// TIA Portal project "CHM_BORDEIRA_20190721" (V15) (continued)
DATA_BLOCK "62_Warning_Data"   // DB62
{ S7_Optimized_Access := 'FALSE' }
VERSION : 0.1
   VAR
      IGG_WARNING_WORD_01 : Word;
      IGG_WARNING_WORD_02 : Word;
      IGG_WARNING_WORD_03 : Word;
      IGG_WARNING_WORD_04 : Word;
      IGG_WARNING_WORD_05 : Word;
      IGG_WARNING_WORD_06 : Word;
      IGG_WARNING_WORD_07 : Word;
      IGG_WARNING_WORD_08 : Word;
      WRNG_PRSNT : Bool;
   END_VAR
BEGIN
END_DATA_BLOCK

DATA_BLOCK "63_E500 Fuel Pumps Not Working_DB"   // DB63
{ S7_Optimized_Access := 'TRUE' }
VERSION : 0.1
// stored: InstanceOfName 63_E500 Fuel Pumps Not Working
"63_E500 Fuel Pumps Not Working"
BEGIN
END_DATA_BLOCK

DATA_BLOCK "64_Message_Data"   // DB64
{ S7_Optimized_Access := 'FALSE' }
VERSION : 0.1
   VAR
      IGG_MESSAGE_WORD_01 : Word;
      IGG_MESSAGE_WORD_02 : Word;
      IGG_MESSAGE_WORD_03 : Word;
      IGG_MESSAGE_WORD_04 : Word;
      IGG_MESSAGE_WORD_05 : Word;
      IGG_MESSAGE_WORD_06 : Word;
      IGG_MESSAGE_WORD_07 : Word;
      IGG_MESSAGE_WORD_08 : Word;
      MSG_PRSNT : Bool;
   END_VAR
BEGIN
END_DATA_BLOCK

DATA_BLOCK "63_Safety System Interlock_IDB"   // DB65
{ S7_Optimized_Access := 'TRUE' }
VERSION : 0.1
// stored: InstanceOfName 64_Safety System Interlock
"64_Safety System Interlock"
BEGIN
END_DATA_BLOCK

DATA_BLOCK "66_Event_Data"   // DB66
{ S7_Optimized_Access := 'FALSE' }
VERSION : 0.1
   VAR
      IGG_EVENT_WORD_01 : Word;
      IGG_EVENT_WORD_02 : Word;
      IGG_EVENT_WORD_03 : Word;
      IGG_EVENT_WORD_04 : Word;
      IGG_EVENT_WORD_05 : Word;
      IGG_EVENT_WORD_06 : Word;
      IGG_EVENT_WORD_07 : Word;
      IGG_EVENT_WORD_08 : Word;
      EVENT_PRSNT : Bool;
   END_VAR
BEGIN
END_DATA_BLOCK

DATA_BLOCK "Alarms_Acknowledge"   // DB67
{ S7_Optimized_Access := 'FALSE' }
VERSION : 0.1
   VAR
      IGG_ALARM_ACKNLG_1 : Word;
      IGG_ALARM_ACKNLG_2 : Word;
      IGG_ALARM_ACKNLG_3 : Word;
      IGG_ALARM_ACKNLG_4 : Word;
      IGG_ALARM_ACKNLG_5 : Word;
      IGG_ALARM_ACKNLG_6 : Word;
   END_VAR
BEGIN
END_DATA_BLOCK

DATA_BLOCK "68_Sys_Status_Data"   // DB68
TITLE = System Status Data
{ S7_Optimized_Access := 'TRUE' }
AUTHOR : JRS
VERSION : 0.1
// Data area for system status information as required by the code
   VAR
      VLVS_AT_INIT : Bool;   // All valves at initial position
      INTRLKS_OK : Bool;   // System interlocks ok
      IA_PRES_IN_RNG : Bool;   // IA Pressure Within Range - PIT112
      CSW_IL_PRES_IN_RNG : Bool;   // CSW Inlet pressure within range - PIT359
      FUEL_PRES_IN_RNG : Bool;   // Fuel pressure within range - PIT204
      OP_PRES_IN_RNG : Bool;   // Output pressure within range - PIT402
      CRG_BLNK_MODE : Bool;   // 1 = Cargon blanketing mode, 0 = Not
      "LOG IGG" : Bool;   // Tag for logging IGG signals
      "STOP LOG IGG" : Bool;
      "LOG IGG Simulator" : Bool;
      "TRUE for HMI" : Bool;
      "E139_SET_SPEED Aux" : Real;
      "E139_SET_SPEED Aux Bool" : Bool;
      "CSW OVR Stop Latched" : Bool;
      "CSW Puls" : Bool;
      "STL Puls" : Bool;
   END_VAR
BEGIN
END_DATA_BLOCK

DATA_BLOCK "503_WARNING CHCK_IDB"   // DB69
{ S7_Optimized_Access := 'TRUE' }
VERSION : 0.1
// stored: InstanceOfName 503_ALARM CHCK
"503_ALARM CHCK"
BEGIN
END_DATA_BLOCK

DATA_BLOCK "CSW_Animation_DB"   // DB71
{ S7_Optimized_Access := 'TRUE' }
VERSION : 0.1
// stored: InstanceOfName Animation
"Animation"
BEGIN
END_DATA_BLOCK

DATA_BLOCK "Ful Pump Ani Animation_DB"   // DB72
{ S7_Optimized_Access := 'TRUE' }
VERSION : 0.1
// stored: InstanceOfName Animation
"Animation"
BEGIN
END_DATA_BLOCK

DATA_BLOCK "IDB_E139"   // DB139
{ S7_Optimized_Access := 'TRUE' }
VERSION : 0.1
// stored: InstanceOfName Animation
"Animation"
BEGIN
END_DATA_BLOCK

DATA_BLOCK "IDB_E500A_Animation"   // DB500
{ S7_Optimized_Access := 'TRUE' }
VERSION : 0.1
// stored: InstanceOfName Animation
"Animation"
BEGIN
END_DATA_BLOCK

DATA_BLOCK "IDB_E500B_Animation"   // DB501
{ S7_Optimized_Access := 'TRUE' }
VERSION : 0.1
// stored: InstanceOfName Animation
"Animation"
BEGIN
END_DATA_BLOCK

DATA_BLOCK "64_Functioning Hours_E500A_IDB"   // DB502
{ S7_Optimized_Access := 'TRUE' }
VERSION : 0.1
// stored: InstanceOfName 64_Functioning Hours
"64_Functioning Hours"
BEGIN
END_DATA_BLOCK

DATA_BLOCK "64_Functioning Hours_E500B_IDB"   // DB503
{ S7_Optimized_Access := 'TRUE' }
VERSION : 0.1
// stored: InstanceOfName 64_Functioning Hours
"64_Functioning Hours"
BEGIN
END_DATA_BLOCK

DATA_BLOCK "Operation hours E139_IDB"   // DB707
{ S7_Optimized_Access := 'TRUE' }
VERSION : 0.1
// stored: InstanceOfName 64_Functioning Hours
"64_Functioning Hours"
BEGIN
END_DATA_BLOCK

DATA_BLOCK "IDB_TIT 315"   // DB715
{ S7_Optimized_Access := 'FALSE' }
VERSION : 0.1
// stored: InstanceOfName 502_ALM_ANALOG
"502_ALM_ANALOG"
BEGIN
END_DATA_BLOCK

DATA_BLOCK "IDB_PIT 316"   // DB716
{ S7_Optimized_Access := 'FALSE' }
VERSION : 0.1
// stored: InstanceOfName 502_ALM_ANALOG
"502_ALM_ANALOG"
BEGIN
END_DATA_BLOCK

DATA_BLOCK "IDB_TIT 319"   // DB719
{ S7_Optimized_Access := 'FALSE' }
VERSION : 0.1
// stored: InstanceOfName 502_ALM_ANALOG
"502_ALM_ANALOG"
BEGIN
END_DATA_BLOCK

DATA_BLOCK "IDB_PIT 102"   // DB722
{ S7_Optimized_Access := 'FALSE' }
VERSION : 0.1
// stored: InstanceOfName 502_ALM_ANALOG
"502_ALM_ANALOG"
BEGIN
END_DATA_BLOCK

DATA_BLOCK "IDB_ATO2B_1"   // DB731
{ S7_Optimized_Access := 'FALSE' }
VERSION : 0.1
// stored: InstanceOfName 502_ALM_ANALOG
"502_ALM_ANALOG"
BEGIN
END_DATA_BLOCK

DATA_BLOCK "IDB_ATO2B_2"   // DB732
{ S7_Optimized_Access := 'FALSE' }
VERSION : 0.1
// stored: InstanceOfName 502_ALM_ANALOG
"502_ALM_ANALOG"
BEGIN
END_DATA_BLOCK

DATA_BLOCK "IDB_TIT 401"   // DB741
{ S7_Optimized_Access := 'FALSE' }
VERSION : 0.1
// stored: InstanceOfName 502_ALM_ANALOG
"502_ALM_ANALOG"
BEGIN
END_DATA_BLOCK

DATA_BLOCK "IDB_PIT 402"   // DB742
{ S7_Optimized_Access := 'FALSE' }
VERSION : 0.1
// stored: InstanceOfName 502_ALM_ANALOG
"502_ALM_ANALOG"
BEGIN
END_DATA_BLOCK

DATA_BLOCK "IDB_PIT 359"   // DB759
{ S7_Optimized_Access := 'FALSE' }
VERSION : 0.1
// stored: InstanceOfName 502_ALM_ANALOG
"502_ALM_ANALOG"
BEGIN
END_DATA_BLOCK

DATA_BLOCK "IDB_TIT 360"   // DB760
{ S7_Optimized_Access := 'FALSE' }
VERSION : 0.1
// stored: InstanceOfName 502_ALM_ANALOG
"502_ALM_ANALOG"
BEGIN
END_DATA_BLOCK

// folder: 70 - 79 Modes of Operation

DATA_BLOCK "70_Mode_Data"   // DB70
{ S7_Optimized_Access := 'TRUE' }
VERSION : 0.1
   VAR
      CRNT_MODE : Int := 1;   // 1 = Auto, 2 = Man, 3 = FatAuto, 4 = FatMan
      INTO_AUTO : Bool;   // Transition to auto
      IN_MAN : Bool;   // In manual
      INTO_AUT_PLS : Bool;   // Pulse bit
      AUT_RST_PLS : TP_TIME;   // Automatic sequence reset pulse
   END_VAR
BEGIN
   AUT_RST_PLS.PT := T#1s;
END_DATA_BLOCK

// folder: 700 - 999 FB Instance DBs

DATA_BLOCK "700_VLV_CHK_DB"   // DB700
{ S7_Optimized_Access := 'TRUE' }
AUTHOR : JRS
VERSION : 0.1
// stored: InstanceOfName 501_VLV_CHK
"501_VLV_CHK"
BEGIN
END_DATA_BLOCK

DATA_BLOCK "701_VLV_CHK_DB"   // DB701
{ S7_Optimized_Access := 'TRUE' }
AUTHOR : JRS
VERSION : 0.1
// stored: InstanceOfName 501_VLV_CHK
"501_VLV_CHK"
BEGIN
END_DATA_BLOCK

DATA_BLOCK "702_VLV_CHK_DB"   // DB702
{ S7_Optimized_Access := 'TRUE' }
AUTHOR : JRS
VERSION : 0.1
// stored: InstanceOfName 501_VLV_CHK
"501_VLV_CHK"
BEGIN
END_DATA_BLOCK

DATA_BLOCK "703_VLV_CHK_DB"   // DB703
{ S7_Optimized_Access := 'TRUE' }
AUTHOR : JRS
VERSION : 0.1
// stored: InstanceOfName 501_VLV_CHK
"501_VLV_CHK"
BEGIN
END_DATA_BLOCK

DATA_BLOCK "704_VLV_CHK_DB"   // DB704
{ S7_Optimized_Access := 'TRUE' }
AUTHOR : JRS
VERSION : 0.1
// stored: InstanceOfName 501_VLV_CHK
"501_VLV_CHK"
BEGIN
END_DATA_BLOCK

DATA_BLOCK "705_VLV_CHK_DB"   // DB705
{ S7_Optimized_Access := 'TRUE' }
AUTHOR : JRS
VERSION : 0.1
// stored: InstanceOfName 501_VLV_CHK
"501_VLV_CHK"
BEGIN
END_DATA_BLOCK

DATA_BLOCK "706_VLV_CHK_DB"   // DB706
{ S7_Optimized_Access := 'TRUE' }
AUTHOR : JRS
VERSION : 0.1
// stored: InstanceOfName 501_VLV_CHK
"501_VLV_CHK"
BEGIN
END_DATA_BLOCK

// folder: 80 - 89 HMI Handling

DATA_BLOCK "80_From_HMI"   // DB80
{ S7_Optimized_Access := 'TRUE' }
VERSION : 0.1
   VAR
      Request_Manual : Bool := False;   // Pulse from HMI
      Request_Auto : Bool := False;   // Pulse from HMI
      SLNCE_BZR : Bool := False;   // Pulse to silence buzzer
      FAT_Mode : Bool := False;   // Set or Reset in HMI
      RST_AUT_SEQ : Bool;   // Reset automatic sequence
      IGG_STND_ALN : Bool := 0;   // 0 = Part of BWT, 1 = Stand Alone
   END_VAR
   VAR RETAIN
      BWT_BYPASS : Bool := TRUE;   // 0 = BWT Control, 1 = BWT Bypassed
   END_VAR
   VAR
      RUN_IGG : Bool;   // Run IGG Command, 1 = Run, 0 = Not
      STOP_IGG : Bool;   // Stop IGG Command, 1 = Stop, 0 = Not
   END_VAR
   VAR RETAIN
      P301_PRSNT : Bool := FALSE;   // 1 = CSW Pump fitted, 0 = Not
      CV312_PRSNT : Bool := TRUE;   // 1 = Scrubber valve fitted, 0 = Not
      CV431_PRSNT : Bool := TRUE;   // 1 = PGC Feed valve fitted, 0 = Not
      CV432_PRSNT : Bool := TRUE;   // 1 = CB Feed valve fitted, 0 = Not
   END_VAR
   VAR
      SW_DTY_PMP_E500 : Bool := 0;   // Button pulse to change duty fuel pump
      MAX_E500_RT : LTime := LT#365d;   // Maximum fuel pump run time
      RST_E500A_RT : Bool;   // Reset runtime for pump A
      RST_E500B_RT : Bool;   // Reset runtime for pump A
   END_VAR
   VAR RETAIN
      E139_SET_SPEED : Real := 1500.0;   // E139 speed in rpm
   END_VAR
   VAR
      CRG_BLNK_MODE : Bool;   // 1 = Cargon blanketing mode, 0 = Not
      MAN_DQ_0_0 : Bool;   // Q0.0 - Fuel Pump #1 Control (E-500-A)
      MAN_DQ_0_1 : Bool;   // Q0.1 - Fuel Pump #2 Control (E-500-B)
      MAN_DQ_0_2 : Bool;   // Q0.2 - CA Blower Control (E139)
      MAN_DQ_0_3 : Bool;   // Q0.3 - Cooling Sea Water (CSW) Inlet Valves Control
      MAN_DQ_0_4 : Bool;   // Q0.4 - Cooling Sea Water (CSW) Outlet Valves Control
      MAN_DQ_0_5 : Bool;   // Q0.5 - IG Supply Valve Control (CV-401)
      MAN_DQ_0_6 : Bool;   // Q0.6 - Cargo Blanketing/BWTS Valve Control (CV431/432)
      MAN_DQ_0_7 : Bool;   // Q0.7 - Spare Output
      MAN_DQ_1_0 : Bool;   // Q1.0 - Spare Output
      MAN_DQ_1_1 : Bool;   // Q1.1 - Atmospheric Alarm (24K2)
      MAN_DQ_1_2 : Bool;   // Q1.2 - IGG Shutdown Alarm Active (24K3)
      MAN_DQ_1_3 : Bool;   // Q1.3 - IGG Warning Alarm Active (24K4)
      MAN_DQ_1_4 : Bool;   // Q1.4 - IGG Running (24PF1)
      MAN_DQ_1_5 : Bool;   // Q1.5 - Shutdown Alarm Active (24PF2)
      MAN_DQ_1_6 : Bool;   // Q1.6 - Warning Alarm Active (24PF3)
      MAN_DQ_1_7 : Bool;   // Q1.7 - Buzzer (24PF4)
      MAN_AQ_INC_98 : Bool;   // QW98 - CV403 - Increase % Signal
      MAN_AQ_DEC_98 : Bool;   // QW98 - CV403 - Decrease % Signal
      MAN_AQ_INC_100 : Bool;   // QW100 - E139 - Increase % Signal
      MAN_AQ_DEC_100 : Bool;   // QW100 - E139 - Decrease % Signal
      MAN_AQ_INC_102 : Bool;   // QW102 - Spare - Increase % Signal
      MAN_AQ_DEC_102 : Bool;   // QW102 - Spare - Decrease % Signal
      MAN_AQ_INC_104 : Bool;   // QW104 - Spare - Increase % Signal
      MAN_AQ_DEC_104 : Bool;   // QW104 - Spare - Decrease % Signal
      RST_LOCKOUT : Bool;
   END_VAR
   VAR RETAIN
      "Beacon frequency" : Time := T#1S;   // Beacon frequency
      "Buzzer reset time" : Time := T#10M;   // Buzzer reset time
   END_VAR
   VAR
      Reset_Alarms : Bool;   // Reset_Alarms
      "Post Purge Time" : Time;
   END_VAR
   VAR RETAIN
      "Cooling System Overrun" : Time := T#30S;
   END_VAR
   VAR
      "PIT 359 delay" : Time := T#2s;
      "PIT 316 delay" : Time := T#2s;
      "CSW OVR Stop" : Bool;   // Puls
   END_VAR
BEGIN
END_DATA_BLOCK

DATA_BLOCK "82_To_HMI"   // DB82
{ S7_Optimized_Access := 'TRUE' }
VERSION : 0.1
   VAR
      CRNT_MODE_IGG : Int := 1;   // 1 = Man, 2 = Auto, 3 = FAT Man, 4 = FATAuto
      "Run Time A" : LTime;   // Run time for pump A
      "Run Time B" : LTime;   // Run time for pump B
      "Duty Is A" : Bool;   // 1 = Duty, 0 = Not
      "Duty Is B" : Bool;   // 1 = Duty, 0 = Not
   END_VAR
   VAR RETAIN
      "CA Blower Run Days" : Int;
      "CA Blower Run Hours" : Int;
      "CA Blower Run Minutes" : Int;
      "CA Blower Run Seconds" : Int;
   END_VAR
   VAR
      "CA Blower Reset Hours" : Bool;
   END_VAR
   VAR RETAIN
      "CA Blower Total Run Hours" : Int;
   END_VAR
   VAR
      "CA Blower Service Due" : Bool;
   END_VAR
   VAR RETAIN
      "CA Blower Service Time Hours" : Int;
      "CA Blower Service Time Days" : Int;
      "CA Blower Hours to Service" : Int;
   END_VAR
   VAR
      "CA Blower Animation" : Int;
      "Fuel Pump 1 Animation" : Int;
      "Fuel Pump 2 Animation" : Int;
   END_VAR
   VAR RETAIN
      "E500A Fuel Pump Run Days" : Int;
      "E500A Fuel Pump Run Hours" : Int;
      "E500A Fuel Pump Run Minutes" : Int;
      "E500A Fuel Pump Run Seconds" : Int;
   END_VAR
   VAR
      "E500A Fuel Pump Reset Hours" : Bool;
   END_VAR
   VAR RETAIN
      "E500A Fuel Pump Total Run Hours" : Int;
   END_VAR
   VAR
      "E500A Fuel Pump Service Due" : Bool;
   END_VAR
   VAR RETAIN
      "E500A Fuel Pump Service Time Hours" : Int;
      "E500A Fuel Pump Service Time Days" : Int;
      "E500A Fuel Pump Hours to Service" : Int;
   END_VAR
   VAR
      "E500A Fuel Pump Animation" : Int;
   END_VAR
   VAR RETAIN
      "E500B Fuel Pump Run Days" : Int;
      "E500B Fuel Pump Run Hours" : Int;
      "E500B Fuel Pump Run Minutes" : Int;
      "E500B Fuel Pump Run Seconds" : Int;
   END_VAR
   VAR
      "E500B Fuel Pump Reset Hours" : Bool;
   END_VAR
   VAR RETAIN
      "E500B Fuel Pump Total Run Hours" : Int;
   END_VAR
   VAR
      "E500B Fuel Pump Service Due" : Bool;
   END_VAR
   VAR RETAIN
      "E500B Fuel Pump Service Time Hours" : Int;
      "E500B Fuel Pump Service Time Days" : Int;
      "E500B Fuel Pump Hours to Service" : Int;
   END_VAR
   VAR
      "E500B Fuel Pump Animation" : Int;
      "IGG RUN Indication" : Bool;
   END_VAR
BEGIN
END_DATA_BLOCK

DATA_BLOCK "84_Setpoints"   // DB84
{ S7_Optimized_Access := 'TRUE' }
VERSION : 0.1
   VAR RETAIN
      PIT112_LowLow : Real := 9.0;   // PIT112 sensor low low setpoint (bar g)
      PIT112_Low : Real := 10.0;   // PIT112 sensor low setpoint (bar g)
      PIT112_High : Real := 20.0;   // PIT112 sensor high setpoint (bar g)
      PIT112_HighHigh : Real := 22.0;   // PIT112 sensor high high setpoint (bar g)
      PIT102_Pilot_LowLow : Real := 15.0;   // PIT102 pilot burner low low setpoint (bar g)
      PIT102_Pilot_Low : Real := 20.0;   // PIT102 pilot burner low setpoint (bar g)
      PIT102_Pilot_High : Real := 200.0;   // PIT102 pilot burner high setpoint (bar g)
      PIT102_Pilot_HighHigh : Real := 300.0;   // PIT102 pilot burner high high setpoint (bar g)
      PIT102_Main_LowLow : Real := 15.0;   // PIT102 main ignition low low setpoint (bar g)
      PIT102_Main_Low : Real := 20.0;   // PIT102 main ignition low setpoint (bar g)
      PIT102_Main_High : Real := 250.0;   // PIT102 main ignition high setpoint (bar g)
      PIT102_Main_HighHigh : Real := 300.0;   // PIT102 main ignition high high setpoint (bar g)
      PIT102_Post_LowLow : Real := 10.0;   // PIT102 post ramp up low low setpoint (bar g)
      PIT102_Post_Low : Real := 15.0;   // PIT102 post ramp up low setpoint (bar g)
      PIT102_Post_High : Real := 250.0;   // PIT102 post ramp up high setpoint (bar g)
      PIT102_Post_HighHigh : Real := 300.0;   // PIT102 post ramp up high high setpoint (bar g)
      PIT204_LowLow : Real := 7.5;   // PIT204 sensor low low setpoint (bar g)
      PIT204_Low : Real := 8.0;   // PIT204 sensor low setpoint (bar g)
      PIT204_High : Real := 11.5;   // PIT204 sensor high setpoint (bar g)
      PIT204_HighHigh : Real := 12.0;   // PIT204 sensor high high setpoint (bar g)
      PIT316_LowLow : Real := 0.1;   // PIT316 sensor low low setpoint (bar g)
      PIT316_Low : Real := 0.2;   // PIT316 sensor low setpoint (bar g)
      PIT316_High : Real := 1.2;   // PIT316 sensor high setpoint (bar g)
      PIT316_HighHigh : Real := 1.4;   // PIT316 sensor high high setpoint (bar g)
      PIT359_LowLow : Real := 0.1;   // PIT359 sensor low low setpoint (bar g)
      PIT359_Low : Real := 0.2;   // PIT359 sensor low setpoint (bar g)
      PIT359_High : Real := 3.0;   // PIT359 sensor high setpoint (bar g)
      PIT359_HighHigh : Real := 3.3;   // PIT359 sensor high high setpoint (bar g)
      PIT402_Pilot_Target : Real := 30.0;   // PIT402 pilot burner target setpoint (bar g)
      PIT402_Pilot_LowLow : Real := 5.0;   // PIT402 pilot burner low low setpoint (bar g)
      PIT402_Pilot_Low : Real := 10.0;   // PIT402 pilot burner low setpoint (bar g)
      PIT402_Pilot_High : Real := 130.0;   // PIT402 pilot burner high setpoint (bar g)
      PIT402_Pilot_HighHigh : Real := 140.0;   // PIT402 pilot burner high high setpoint (bar g)
      PIT402_Main_Target : Real := 40.0;   // PIT402 main ignirition target setpoint (bar g)
      PIT402_Main_LowLow : Real := 5.0;   // PIT402 main ignirition low low setpoint (bar g)
      PIT402_Main_Low : Real := 10.0;   // PIT402 main ignirition low setpoint (bar g)
      PIT402_Main_High : Real := 250.0;   // PIT402 main ignirition high setpoint (bar g)
      PIT402_Main_HighHigh : Real := 300.0;   // PIT402 main ignirition high high setpoint (bar g)
      PIT402_Post_Target_Start : Real := 50.0;   // PIT402 post ramp up target start setpoint (bar g)
      PIT401_Post_Target_Max : Real := 150.0;   // PIT402 post ramp up target max setpoint (bar g)
      PIT402_Post_LowLow : Real := 5.0;   // PIT402 post ramp up low low setpoint (bar g)
      PIT402_Post_Low : Real := 10.0;   // PIT402 post ramp up low setpoint (bar g)
      PIT402_Post_High : Real := 250.0;   // PIT402 post ramp up high setpoint (bar g)
      PIT402_Post_HighHigh : Real := 300.0;   // PIT402 post ramp up high high setpoint (bar g)
      TIT315_High : Real := 47.0;   // TIT315 sensor high setpoint (degC)
      TIT315_HighHigh : Real := 50.0;   // TIT315 sensor high high setpoint (degC)
      TIT319_High : Real := 37.0;   // TIT319 sensor high setpoint (degC)
      TIT319_HighHigh : Real := 40.0;   // TIT319 sensor high high setpoint (degC)
      TIT360_High : Real := 47.0;   // TIT360 sensor high setpoint (degC)
      TIT360_HighHigh : Real := 50.0;   // TIT360 sensor high high setpoint (degC)
      TIT401_High : Real := 50.0;   // TIT401 sensor high setpoint (degC)
      TIT401_HighHigh : Real := 55.5;   // TIT401 sensor high high setpoint (degC)
      AT_O2_1_LowLow : Real := 18.5;   // Atmospheric O2 sensor #1 LowLow setpoint
      AT_O2_1_Low : Real := 19.0;   // Atmospheric O2 sensor #1 Low setpoint
      AT_O2_2_LowLow : Real := 18.5;   // Atmospheric O2 sensor #2 LowLow setpoint
      AT_O2_2_Low : Real := 19.0;   // Atmospheric O2 sensor #2 Low setpoint
   END_VAR
BEGIN
END_DATA_BLOCK

DATA_BLOCK "86_Times"   // DB86
{ S7_Optimized_Access := 'TRUE' }
VERSION : 0.1
   VAR RETAIN
      PRE_BC_STRT_CMND_DLY : Time := T#5S;   // Time delay prior to IGG to BC start command
      PRE_CV203_CLS_CMND_DLY : Time := T#3S;   // Time delay prior to CV203 close command
      POST_P301_STOP_DLY : Time := T#1S;   // Time delay after P301 stopped
      POST_CV311_CLS_DLY : Time := T#3S;   // Time delay after CV311 closed (CV312 opened)
      POST_CV321_OPN_DLY : Time := T#3S;   // Time delay after CV321 opened (CV322 closed)
      CV311_MAX_TRVL_TIME : Time := T#30S;   // Maximum valve travel time
      CV312_MAX_TRVL_TIME : Time := T#30S;   // Maximum valve travel time
      CV321_MAX_TRVL_TIME : Time := T#2M;   // Maximum valve travel time
      CV322_MAX_TRVL_TIME : Time := T#1M;   // Maximum valve travel time
      CV401_MAX_TRVL_TIME : Time := T#30S;   // Maximum valve travel time
      CV431_MAX_TRVL_TIME : Time := T#30S;   // Maximum valve travel time
      CV432_MAX_TRVL_TIME : Time := T#30S;   // Maximum valve travel time
      PIT402_Ramp_Seconds : Int := 30;   // Time in seconds for target ramp up
   END_VAR
   VAR
      STEP_MAX_TIME_STP_001 : Time := T#5S;
      STEP_MAX_TIME_STP_005 : Time := T#5S;
      STEP_MAX_TIME_STP_010 : Time := T#5S;
      STEP_MAX_TIME_STP_020 : Time := T#5S;
      STEP_MAX_TIME_STP_030 : Time := T#5S;
      STEP_MAX_TIME_STP_040 : Time := T#5S;
      STEP_MAX_TIME_STP_050 : Time := T#5S;
      STEP_MAX_TIME_STP_060 : Time := T#5S;
      STEP_MAX_TIME_STP_070 : Time := T#5S;
      STEP_MAX_TIME_STP_080 : Time := T#5S;
      STEP_MAX_TIME_STP_090 : Time := T#5S;
      STEP_MAX_TIME_STP_100 : Time := T#30S;
      STEP_MAX_TIME_STP_110 : Time := T#5S;
      STEP_MAX_TIME_STP_120 : Time := T#5S;
      STEP_MAX_TIME_STP_130 : Time := T#5S;
      STEP_MAX_TIME_STP_140 : Time := T#5S;
      STEP_MAX_TIME_STP_150 : Time := T#5S;
      STEP_MAX_TIME_STP_160 : Time := T#5S;
      STEP_MAX_TIME_STP_170 : Time := T#5S;
      STEP_MAX_TIME_STP_180 : Time := T#5S;
      STEP_MAX_TIME_STP_190 : Time := T#5S;
      STEP_MAX_TIME_STP_200 : Time := T#5S;
      STEP_MAX_TIME_STP_210 : Time := T#5S;
      STEP_MAX_TIME_STP_220 : Time := T#5S;
      STEP_MAX_TIME_STP_230 : Time := T#5S;
      STEP_MAX_TIME_STP_240 : Time := T#5S;
      STEP_MAX_TIME_STP_250 : Time := T#5S;
      STEP_MAX_TIME_STP_260 : Time := T#5S;
      STEP_MAX_TIME_STP_270 : Time := T#5S;
      STEP_MAX_TIME_STP_280 : Time := T#5S;
      STEP_MAX_TIME_STP_290 : Time := T#5S;
      STEP_MAX_TIME_STP_300 : Time := T#5S;
      STEP_MAX_TIME_STP_310 : Time := T#5S;
      STEP_MAX_TIME_STP_320 : Time := T#5S;
      STEP_MAX_TIME_STP_330 : Time := T#5S;
      STEP_MAX_TIME_STP_340 : Time := T#5S;
      STEP_MAX_TIME_STP_350 : Time := T#5S;
      STEP_MAX_TIME_STP_360 : Time := T#5S;
      STEP_MAX_TIME_STP_370 : Time := T#5S;
      STEP_MAX_TIME_STP_380 : Time := T#30S;
      STEP_MAX_TIME_STP_390 : Time := T#5S;
      STEP_MAX_TIME_STP_400 : Time := T#5S;
      STEP_MAX_TIME_STP_410 : Time := T#5S;
      STEP_MAX_TIME_STP_420 : Time := T#5S;
      STEP_MAX_TIME_STP_430 : Time := T#5S;
      STEP_MAX_TIME_STP_440 : Time := T#5S;
      STEP_MAX_TIME_STP_450 : Time := T#5S;
      STEP_MAX_TIME_STP_460 : Time := T#5S;
      STEP_MAX_TIME_STP_470 : Time := T#5S;
      STEP_MAX_TIME_STP_480 : Time := T#5S;
      STEP_MAX_TIME_STP_490 : Time := T#5S;
      STEP_MAX_TIME_STP_500 : Time := T#5S;
   END_VAR
   VAR RETAIN
      "PIT402 Alarm Delay" : Time := T#2M;
   END_VAR
BEGIN
END_DATA_BLOCK

// folder: 90 - 99 Manual Functions

DATA_BLOCK "90_Manual_Data"   // DB90
{ S7_Optimized_Access := 'TRUE' }
VERSION : 0.1
   VAR
      INC_PLS_98 : Bool;   // Pulse bit
      INC_PLS_98_Hz : Bool;   // Pulse bit
      DEC_PLS_98 : Bool;   // Pulse bit
      DEC_PLS_98_Hz : Bool;   // Pulse bit
      INC_PLS_100 : Bool;   // Pulse bit
      INC_PLS_100_Hz : Bool;   // Pulse bit
      DEC_PLS_100 : Bool;   // Pulse bit
      DEC_PLS_100_Hz : Bool;   // Pulse bit
      INC_PLS_102 : Bool;   // Pulse bit
      INC_PLS_102_Hz : Bool;   // Pulse bit
      DEC_PLS_102 : Bool;   // Pulse bit
      DEC_PLS_102_Hz : Bool;   // Pulse bit
      INC_PLS_104 : Bool;   // Pulse bit
      INC_PLS_104_Hz : Bool;   // Pulse bit
      DEC_PLS_104 : Bool;   // Pulse bit
      DEC_PLS_104_Hz : Bool;   // Pulse bit
   END_VAR
BEGIN
END_DATA_BLOCK

DATA_BLOCK "E500A"   // DB505
{ S7_Optimized_Access := 'TRUE' }
VERSION : 0.1
// stored: InstanceOfName FuelPump
"FuelPump"
BEGIN
END_DATA_BLOCK

// folder: System blocks/Program resources

DATA_BLOCK "TON Delay Low IG Pressure"   // DB22
{ S7_Optimized_Access := 'TRUE' }
AUTHOR : Simatic
FAMILY : IEC
NAME : IEC_TMR
VERSION : 1.0
// stored: InstanceOfName IEC_TIMER
"IEC_TIMER"
BEGIN
END_DATA_BLOCK

// folder: (top level)

ORGANIZATION_BLOCK "IGG Main PLC"   // OB1, LAD, ProgramCycle
TITLE = "Main Program Sweep (Cycle)"
{ S7_Optimized_Access := 'TRUE' }
VERSION : 0.1
   VAR_INPUT
      Initial_Call : Bool;   // Initial call of this OB
      Remanence : Bool;   // =True, if remanent data are available
   END_VAR
   VAR_TEMP   // added for the SCL form of the ladder/FBD networks
      _w1 : Bool;
   END_VAR
BEGIN

REGION Network 1: Digital Input Processing
   // To process raw inputs prior to code use
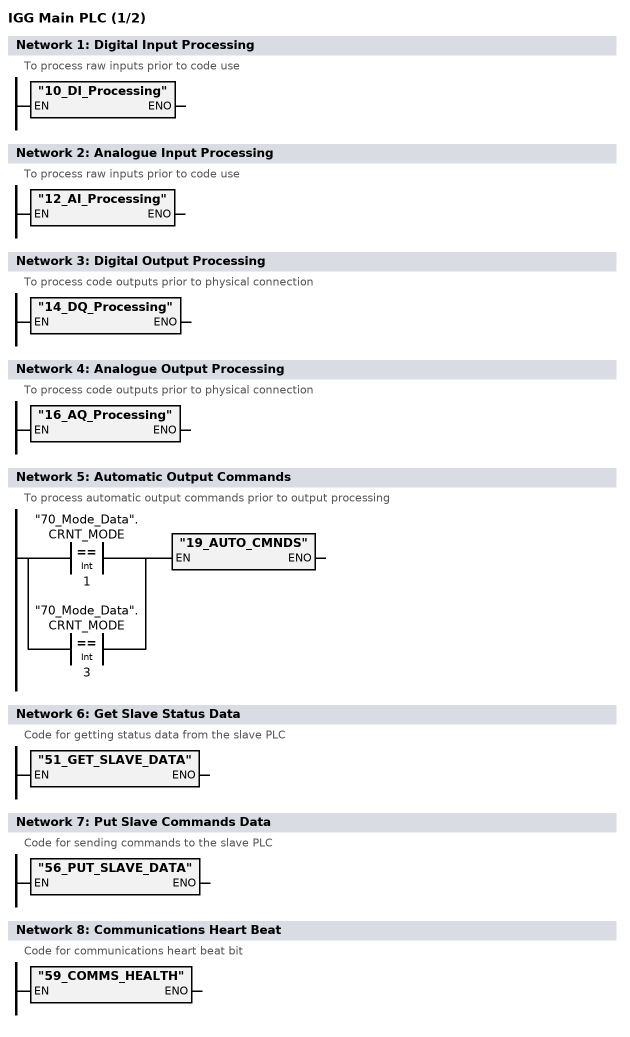
   RUNG wire#powerrail
      "10_DI_Processing"()
   END_RUNG
   // the same network as SCL:
   "10_DI_Processing"();
END_REGION

REGION Network 2: Analogue Input Processing
   // To process raw inputs prior to code use
   RUNG wire#powerrail
      "12_AI_Processing"()
   END_RUNG
   // the same network as SCL:
   "12_AI_Processing"();
END_REGION

REGION Network 3: Digital Output Processing
   // To process code outputs prior to physical connection
   RUNG wire#powerrail
      "14_DQ_Processing"()
   END_RUNG
   // the same network as SCL:
   "14_DQ_Processing"();
END_REGION

REGION Network 4: Analogue Output Processing
   // To process code outputs prior to physical connection
   RUNG wire#powerrail
      "16_AQ_Processing"()
   END_RUNG
   // the same network as SCL:
   "16_AQ_Processing"();
END_REGION

REGION Network 5: Automatic Output Commands
   // To process automatic output commands prior to output processing
   RUNG wire#powerrail
      { S7_Templates := "SrcType := Int" } EQ_Contact(in1 := "70_Mode_Data".CRNT_MODE, in2 := 1)
      wire#w1
      "19_AUTO_CMNDS"()
   END_RUNG
   RUNG wire#powerrail
      { S7_Templates := "SrcType := Int" } EQ_Contact(in1 := "70_Mode_Data".CRNT_MODE, in2 := 3)
   END_RUNG wire#w1
   // the same network as SCL:
   IF ("70_Mode_Data".CRNT_MODE = 1) OR ("70_Mode_Data".CRNT_MODE = 3) THEN "19_AUTO_CMNDS"(); END_IF;
END_REGION

REGION Network 6: Get Slave Status Data
   // Code for getting status data from the slave PLC
   RUNG wire#powerrail
      "51_GET_SLAVE_DATA"()
   END_RUNG
   // the same network as SCL:
   "51_GET_SLAVE_DATA"();
END_REGION

REGION Network 7: Put Slave Commands Data
   // Code for sending commands to the slave PLC
   RUNG wire#powerrail
      "56_PUT_SLAVE_DATA"()
   END_RUNG
   // the same network as SCL:
   "56_PUT_SLAVE_DATA"();
END_REGION

REGION Network 8: Communications Heart Beat
   // Code for communications heart beat bit
   RUNG wire#powerrail
      "59_COMMS_HEALTH"()
   END_RUNG
   // the same network as SCL:
   "59_COMMS_HEALTH"();
END_REGION

REGION Network 9: Alarm Handling
   // Code to determine alarm conditions
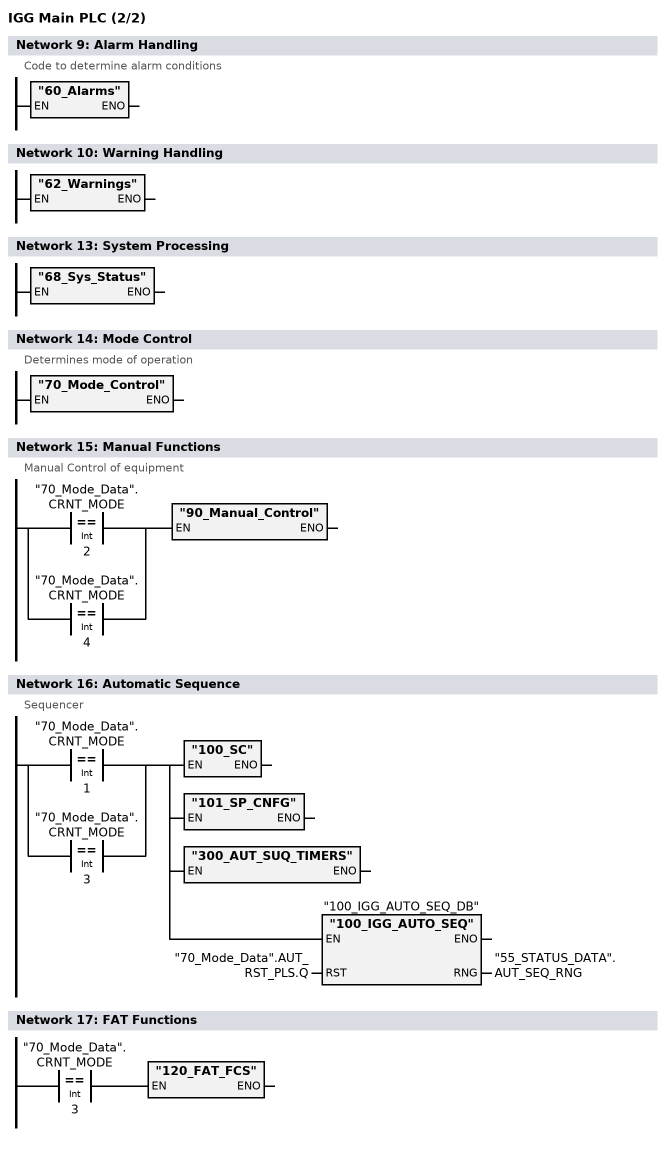
   RUNG wire#powerrail
      "60_Alarms"()
   END_RUNG
   // the same network as SCL:
   "60_Alarms"();
END_REGION

REGION Network 10: Warning Handling
   RUNG wire#powerrail
      "62_Warnings"()
   END_RUNG
   // the same network as SCL:
   "62_Warnings"();
END_REGION

REGION Network 11: Message Handling
   // Handles messaging
END_REGION

REGION Network 12: Event Handling
   // Records event data
END_REGION

REGION Network 13: System Processing
   RUNG wire#powerrail
      "68_Sys_Status"()
   END_RUNG
   // the same network as SCL:
   "68_Sys_Status"();
END_REGION

REGION Network 14: Mode Control
   // Determines mode of operation
   RUNG wire#powerrail
      "70_Mode_Control"()
   END_RUNG
   // the same network as SCL:
   "70_Mode_Control"();
END_REGION

REGION Network 15: Manual Functions
   // Manual Control of equipment
   RUNG wire#powerrail
      { S7_Templates := "SrcType := Int" } EQ_Contact(in1 := "70_Mode_Data".CRNT_MODE, in2 := 2)
      wire#w1
      "90_Manual_Control"()
   END_RUNG
   RUNG wire#powerrail
      { S7_Templates := "SrcType := Int" } EQ_Contact(in1 := "70_Mode_Data".CRNT_MODE, in2 := 4)
   END_RUNG wire#w1
   // the same network as SCL:
   IF ("70_Mode_Data".CRNT_MODE = 2) OR ("70_Mode_Data".CRNT_MODE = 4) THEN "90_Manual_Control"(); END_IF;
END_REGION

REGION Network 16: Automatic Sequence
   // Sequencer
   RUNG wire#powerrail
      { S7_Templates := "SrcType := Int" } EQ_Contact(in1 := "70_Mode_Data".CRNT_MODE, in2 := 1)
      wire#w1
      "100_SC"()
   END_RUNG
   RUNG wire#powerrail
      { S7_Templates := "SrcType := Int" } EQ_Contact(in1 := "70_Mode_Data".CRNT_MODE, in2 := 3)
   END_RUNG wire#w1
   RUNG wire#w1
      "101_SP_CNFG"()
   END_RUNG
   RUNG wire#w1
      "300_AUT_SUQ_TIMERS"()
   END_RUNG
   RUNG wire#w1
      "100_IGG_AUTO_SEQ_DB"(RST := "70_Mode_Data".AUT_RST_PLS.Q, RNG => "55_STATUS_DATA".AUT_SEQ_RNG)
   END_RUNG
   // the same network as SCL:
   #_w1 := ("70_Mode_Data".CRNT_MODE = 1) OR ("70_Mode_Data".CRNT_MODE = 3);
   IF #_w1 THEN
       "100_SC"();
       "101_SP_CNFG"();
       "300_AUT_SUQ_TIMERS"();
       "100_IGG_AUTO_SEQ_DB"(RST := "70_Mode_Data".AUT_RST_PLS.Q, RNG => "55_STATUS_DATA".AUT_SEQ_RNG);   // "100_IGG_AUTO_SEQ"
   END_IF;
END_REGION

REGION Network 17: FAT Functions
   RUNG wire#powerrail
      { S7_Templates := "SrcType := Int" } EQ_Contact(in1 := "70_Mode_Data".CRNT_MODE, in2 := 3)
      "120_FAT_FCS"()
   END_RUNG
   // the same network as SCL:
   IF "70_Mode_Data".CRNT_MODE = 3 THEN "120_FAT_FCS"(); END_IF;
END_REGION
END_ORGANIZATION_BLOCK

// folder: 10 - 19 IO & Processing

FUNCTION "10_DI_Processing" : Void   // FC10, LAD
TITLE = Digital Input Processing
{ S7_Optimized_Access := 'TRUE' }
AUTHOR : JRS
VERSION : 0.1
// To process raw inputs prior to code use
BEGIN

REGION Network 1: I0.0 - IGG E-Stop Healthy (S2-8K1)
   // True = OK, False = NOK
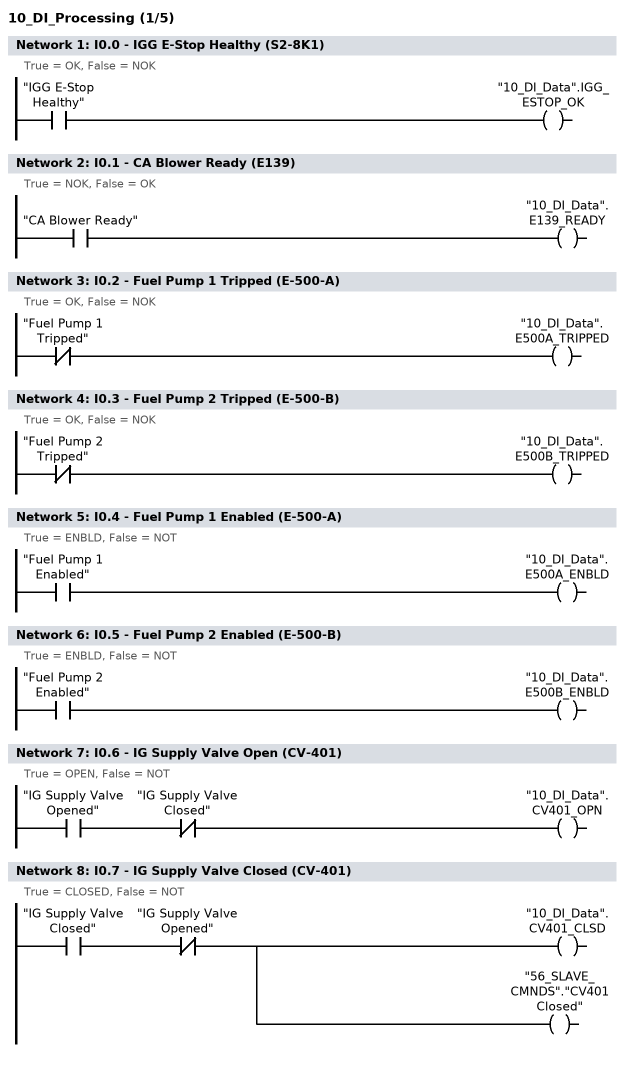
   RUNG wire#powerrail
      Contact( "IGG E-Stop Healthy" )
      Coil( "10_DI_Data".IGG_ESTOP_OK )
   END_RUNG
   // the same network as SCL:
   "10_DI_Data".IGG_ESTOP_OK := "IGG E-Stop Healthy";
END_REGION

REGION Network 2: I0.1 - CA Blower Ready (E139)
   // True = NOK, False = OK
   RUNG wire#powerrail
      Contact( "CA Blower Ready" )
      Coil( "10_DI_Data".E139_READY )
   END_RUNG
   // the same network as SCL:
   "10_DI_Data".E139_READY := "CA Blower Ready";
END_REGION

REGION Network 3: I0.2 - Fuel Pump 1 Tripped (E-500-A)
   // True = OK, False = NOK
   RUNG wire#powerrail
      I_Contact( "Fuel Pump 1 Tripped" )
      Coil( "10_DI_Data".E500A_TRIPPED )
   END_RUNG
   // the same network as SCL:
   "10_DI_Data".E500A_TRIPPED := NOT "Fuel Pump 1 Tripped";
END_REGION

REGION Network 4: I0.3 - Fuel Pump 2 Tripped (E-500-B)
   // True = OK, False = NOK
   RUNG wire#powerrail
      I_Contact( "Fuel Pump 2 Tripped" )
      Coil( "10_DI_Data".E500B_TRIPPED )
   END_RUNG
   // the same network as SCL:
   "10_DI_Data".E500B_TRIPPED := NOT "Fuel Pump 2 Tripped";
END_REGION

REGION Network 5: I0.4 - Fuel Pump 1 Enabled (E-500-A)
   // True = ENBLD, False = NOT
   RUNG wire#powerrail
      Contact( "Fuel Pump 1 Enabled" )
      Coil( "10_DI_Data".E500A_ENBLD )
   END_RUNG
   // the same network as SCL:
   "10_DI_Data".E500A_ENBLD := "Fuel Pump 1 Enabled";
END_REGION

REGION Network 6: I0.5 - Fuel Pump 2 Enabled (E-500-B)
   // True = ENBLD, False = NOT
   RUNG wire#powerrail
      Contact( "Fuel Pump 2 Enabled" )
      Coil( "10_DI_Data".E500B_ENBLD )
   END_RUNG
   // the same network as SCL:
   "10_DI_Data".E500B_ENBLD := "Fuel Pump 2 Enabled";
END_REGION

REGION Network 7: I0.6 - IG Supply Valve Open (CV-401)
   // True = OPEN, False = NOT
   RUNG wire#powerrail
      Contact( "IG Supply Valve Opened" )
      I_Contact( "IG Supply Valve Closed" )
      Coil( "10_DI_Data".CV401_OPN )
   END_RUNG
   // the same network as SCL:
   "10_DI_Data".CV401_OPN := "IG Supply Valve Opened" AND NOT "IG Supply Valve Closed";
END_REGION

REGION Network 8: I0.7 - IG Supply Valve Closed (CV-401)
   // True = CLOSED, False = NOT
   RUNG wire#powerrail
      Contact( "IG Supply Valve Closed" )
      I_Contact( "IG Supply Valve Opened" )
      wire#w1
      Coil( "10_DI_Data".CV401_CLSD )
   END_RUNG
   RUNG wire#w1
      Coil( "56_SLAVE_CMNDS"."CV401 Closed" )
   END_RUNG
   // the same network as SCL:
   "10_DI_Data".CV401_CLSD := "IG Supply Valve Closed" AND NOT "IG Supply Valve Opened";
   "56_SLAVE_CMNDS"."CV401 Closed" := "10_DI_Data".CV401_CLSD;
END_REGION

REGION Network 9: I1.0 - DTB Valve Open (CV-321)
   // True = OPEN, False = NOT
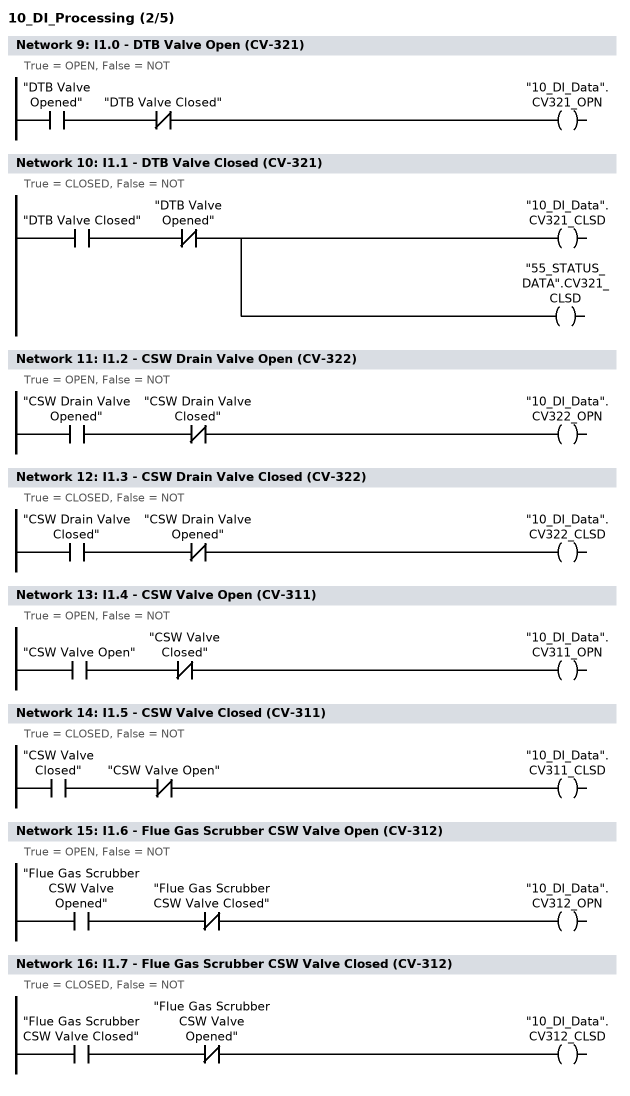
   RUNG wire#powerrail
      Contact( "DTB Valve Opened" )
      I_Contact( "DTB Valve Closed" )
      Coil( "10_DI_Data".CV321_OPN )
   END_RUNG
   // the same network as SCL:
   "10_DI_Data".CV321_OPN := "DTB Valve Opened" AND NOT "DTB Valve Closed";
END_REGION

REGION Network 10: I1.1 - DTB Valve Closed (CV-321)
   // True = CLOSED, False = NOT
   RUNG wire#powerrail
      Contact( "DTB Valve Closed" )
      I_Contact( "DTB Valve Opened" )
      wire#w1
      Coil( "10_DI_Data".CV321_CLSD )
   END_RUNG
   RUNG wire#w1
      Coil( "55_STATUS_DATA".CV321_CLSD )
   END_RUNG
   // the same network as SCL:
   "10_DI_Data".CV321_CLSD := "DTB Valve Closed" AND NOT "DTB Valve Opened";
   "55_STATUS_DATA".CV321_CLSD := "10_DI_Data".CV321_CLSD;
END_REGION

REGION Network 11: I1.2 - CSW Drain Valve Open (CV-322)
   // True = OPEN, False = NOT
   RUNG wire#powerrail
      Contact( "CSW Drain Valve Opened" )
      I_Contact( "CSW Drain Valve Closed" )
      Coil( "10_DI_Data".CV322_OPN )
   END_RUNG
   // the same network as SCL:
   "10_DI_Data".CV322_OPN := "CSW Drain Valve Opened" AND NOT "CSW Drain Valve Closed";
END_REGION

REGION Network 12: I1.3 - CSW Drain Valve Closed (CV-322)
   // True = CLOSED, False = NOT
   RUNG wire#powerrail
      Contact( "CSW Drain Valve Closed" )
      I_Contact( "CSW Drain Valve Opened" )
      Coil( "10_DI_Data".CV322_CLSD )
   END_RUNG
   // the same network as SCL:
   "10_DI_Data".CV322_CLSD := "CSW Drain Valve Closed" AND NOT "CSW Drain Valve Opened";
END_REGION

REGION Network 13: I1.4 - CSW Valve Open (CV-311)
   // True = OPEN, False = NOT
   RUNG wire#powerrail
      Contact( "CSW Valve Open" )
      I_Contact( "CSW Valve Closed" )
      Coil( "10_DI_Data".CV311_OPN )
   END_RUNG
   // the same network as SCL:
   "10_DI_Data".CV311_OPN := "CSW Valve Open" AND NOT "CSW Valve Closed";
END_REGION
